// TIA Portal project "ProjectTest" (V15.1)

(* hardware
DEVICE "S7-1200 station_1"  S7-1200 Station
   slot 0: "Rack_0"  S7-1200 Rack  Rack  V1.0
   slot 1: "PLC_1"  CPU 1214C DC/DC/DC  6ES7 214-1AG40-0XB0  V4.2
DEVICE "HMI_1"  KTP900 Basic PN
   slot 0: "HMI_1"  KTP900 Basic PN  6AV2 123-2JB03-0AX0  15.1.0.0
   slot 1: "HMI_RT_1"  KTP900 Basic PN  6AV2 123-2JB03-0AX0  15.1.0.0
   slot 5: "HMI_1.IE_CP_1"  PROFINET Interface  15.0.1.0
      slot 1: "PROFINET Interface_1"  PROFINET Interface
         slot 1: "Port_1"  Port
*)

// ===== PLC "PLC_1"  CPU 1214C DC/DC/DC =====

VAR_GLOBAL   // PLC tag table "Default tag table"
   "System_Byte" AT %MB1 : Byte;
   "FirstScan" AT %M1.0 : Bool;
   "DiagStatusUpdate" AT %M1.1 : Bool;
   "AlwaysTRUE" AT %M1.2 : Bool;
   "AlwaysFALSE" AT %M1.3 : Bool;
   "Clock_Byte" AT %MB0 : Byte;
   "Clock_10Hz" AT %M0.0 : Bool;
   "Clock_5Hz" AT %M0.1 : Bool;
   "Clock_2.5Hz" AT %M0.2 : Bool;
   "Clock_2Hz" AT %M0.3 : Bool;
   "Clock_1.25Hz" AT %M0.4 : Bool;
   "Clock_1Hz" AT %M0.5 : Bool;
   "Clock_0.625Hz" AT %M0.6 : Bool;
   "Clock_0.5Hz" AT %M0.7 : Bool;
   "puls" AT %M2.0 : Bool;
END_VAR

VAR_GLOBAL   // PLC tag table "Tags_DI"
   "Pompa1" AT %Q0.0 : Bool;
   "Pompa2" AT %Q0.1 : Bool;
   "Vana Consum" AT %Q0.2 : Bool;
   "Buton pompa1" AT %I0.0 : Bool;
   "Buton Pompa2" AT %I0.1 : Bool;
   "Buton Vana" AT %I0.2 : Bool;
   "Resetare Contor1" AT %I0.3 : Bool;
   "Resetare Contor2" AT %I0.4 : Bool;
   "Indicatie Pompa1" AT %I0.5 : Bool;
   "Indicatie Pompa2" AT %I0.6 : Bool;
   "Indicatie mod" AT %I0.7 : Bool;
END_VAR

DATA_BLOCK "Bazin"   // DB1
{ S7_Optimized_Access := 'TRUE' }
VERSION : 0.1
   VAR
      Nivel : Real;
      "Vana golire" : Bool := false;
      "Debit golire" : Int := 10;
      Cheie : Int := 1;
      Stare_rising_edge : Bool;
   END_VAR
BEGIN
END_DATA_BLOCK

DATA_BLOCK "Pompa_1"   // DB2
{ S7_Optimized_Access := 'TRUE' }
VERSION : 0.1
   VAR
      Stare : Bool;
      Capacitate : Real := 15.0;
      "Mod" : Int;
      Contor : UInt;
      Stare_rising_edge_bazin : Bool;
      Reset : Bool;
      add_15l : Real := 15.0;
      Stare_rising_edge_pompa : Bool;
   END_VAR
BEGIN
END_DATA_BLOCK

DATA_BLOCK "Pompa_2"   // DB3
{ S7_Optimized_Access := 'TRUE' }
VERSION : 0.1
   VAR
      Stare : Bool;
      Capacitate : Real := 15.0;
      "Mod" : Int;
      Contor : UInt;
      Stare_rising_edge_bazin : Bool;
      Reset : Bool;
      add_15l : Real := 15.0;
      State_rising_edge_pompa : Bool;
   END_VAR
BEGIN
END_DATA_BLOCK

DATA_BLOCK "Adauga  15L la bazin_DB"   // DB4
{ S7_Optimized_Access := 'TRUE' }
VERSION : 0.1
// stored: InstanceOfName Adauga 15L la bazin
"Adauga  15L la bazin"
BEGIN
END_DATA_BLOCK

DATA_BLOCK "Adauga  15L la bazin_DB_1"   // DB5
{ S7_Optimized_Access := 'TRUE' }
VERSION : 0.1
// stored: InstanceOfName Adauga 15L la bazin
"Adauga  15L la bazin"
BEGIN
END_DATA_BLOCK

DATA_BLOCK "Adauga  15L la bazin_DB_2"   // DB6
{ S7_Optimized_Access := 'TRUE' }
VERSION : 0.1
// stored: InstanceOfName Adauga 15L la bazin
"Adauga  15L la bazin"
BEGIN
END_DATA_BLOCK

DATA_BLOCK "Adauga  15L la bazin_DB_3"   // DB7
{ S7_Optimized_Access := 'TRUE' }
VERSION : 0.1
// stored: InstanceOfName Adauga 15L la bazin
"Adauga  15L la bazin"
BEGIN
END_DATA_BLOCK

DATA_BLOCK "Adauga  15L la bazin_DB_4"   // DB8
{ S7_Optimized_Access := 'TRUE' }
VERSION : 0.1
// stored: InstanceOfName Adauga 15L la bazin
"Adauga  15L la bazin"
BEGIN
END_DATA_BLOCK

DATA_BLOCK "Adauga  15L la bazin_DB_5"   // DB9
{ S7_Optimized_Access := 'TRUE' }
VERSION : 0.1
// stored: InstanceOfName Adauga 15L la bazin
"Adauga  15L la bazin"
BEGIN
END_DATA_BLOCK

FUNCTION_BLOCK "Adauga  15L la bazin"   // FB1, LAD
{ S7_Optimized_Access := 'TRUE' }
VERSION : 0.1
   VAR_INPUT
      Input_2 : Bool;
   END_VAR
   VAR_TEMP
      clock_rising_edge : Bool;
   END_VAR
   VAR_TEMP   // added for the SCL form of the ladder/FBD networks
      _w1 : Bool;
      _w2 : Bool;
   END_VAR
BEGIN

REGION Network 1
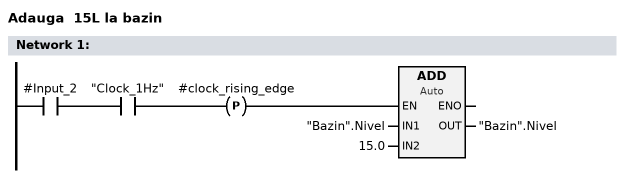
   RUNG wire#powerrail
      Contact( #Input_2 )
      Contact( "Clock_1Hz" )
      P_Trig( #clock_rising_edge )
      Add(in1 := "Bazin".Nivel, in2 := 15.0, out => "Bazin".Nivel)
   END_RUNG
   // the same network as SCL:
   #_w1 := #Input_2 AND "Clock_1Hz";
   #_w2 := #_w1 AND NOT #clock_rising_edge;   // rising edge
   #clock_rising_edge := #_w1;
   IF #_w2 THEN "Bazin".Nivel := "Bazin".Nivel + 15.0; END_IF;
END_REGION
END_FUNCTION_BLOCK

FUNCTION "Block_1" : Void   // FC1, LAD
{ S7_Optimized_Access := 'TRUE' }
VERSION : 0.1
   VAR_INPUT
      input1 : Bool;
   END_VAR
   VAR_TEMP
      clock_rising_edge : Bool;
   END_VAR
   VAR_TEMP   // added for the SCL form of the ladder/FBD networks
      _w1 : Bool;
      _w2 : Bool;
   END_VAR
BEGIN

REGION Network 1
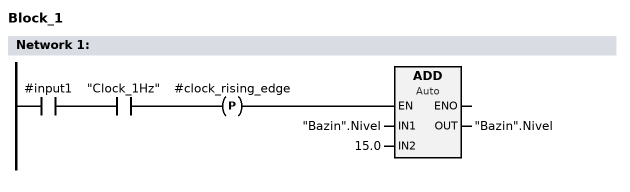
   RUNG wire#powerrail
      Contact( #input1 )
      Contact( "Clock_1Hz" )
      P_Trig( #clock_rising_edge )
      Add(in1 := "Bazin".Nivel, in2 := 15.0, out => "Bazin".Nivel)
   END_RUNG
   // the same network as SCL:
   #_w1 := #input1 AND "Clock_1Hz";
   #_w2 := #_w1 AND NOT #clock_rising_edge;   // rising edge
   #clock_rising_edge := #_w1;
   IF #_w2 THEN "Bazin".Nivel := "Bazin".Nivel + 15.0; END_IF;
END_REGION
END_FUNCTION

ORGANIZATION_BLOCK "Main"   // OB1, LAD, ProgramCycle
TITLE = "Main Program Sweep (Cycle)"
{ S7_Optimized_Access := 'TRUE' }
VERSION : 0.1
   VAR_INPUT
      Initial_Call : Bool;   // Initial call of this OB
      Remanence : Bool;   // =True, if remanent data are available
   END_VAR
   VAR_TEMP   // added for the SCL form of the ladder/FBD networks
      _w1 : Bool;
      _w2 : Bool;
      _w3 : Bool;
      _w4 : Bool;
   END_VAR
BEGIN

REGION Network 1: moduri de functionare
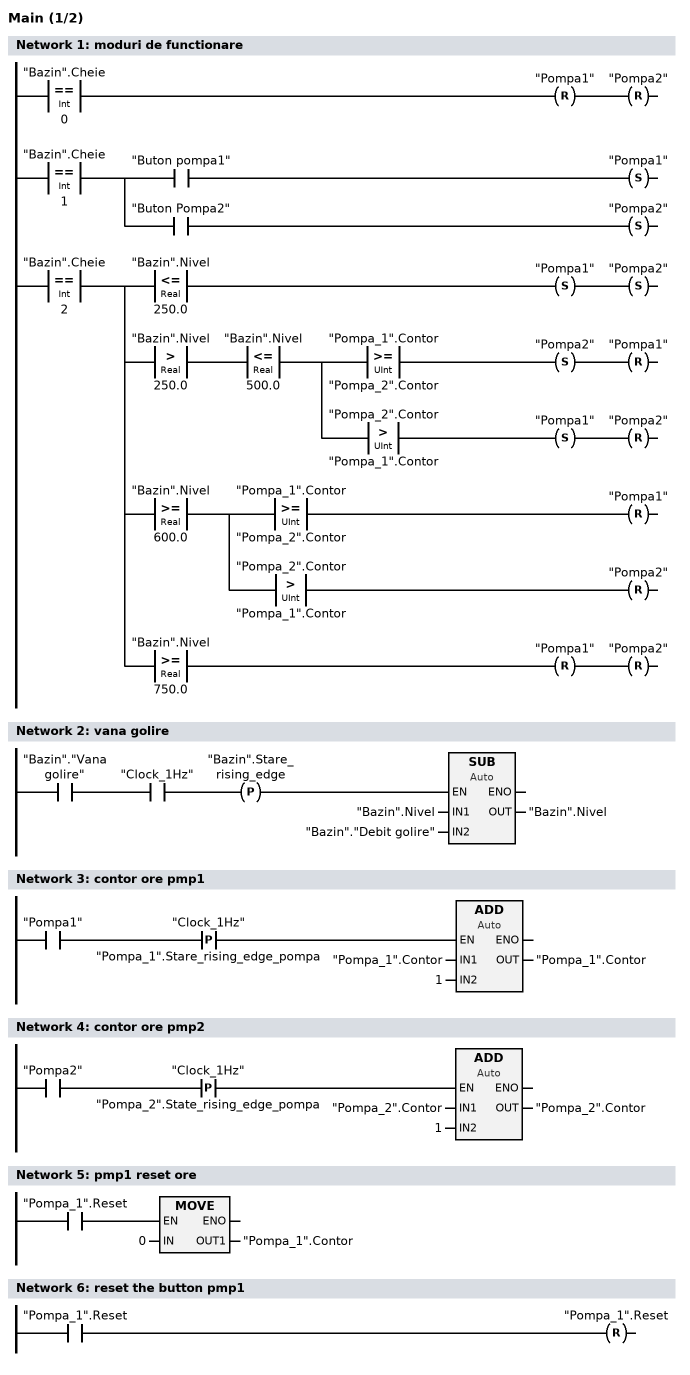
   RUNG wire#powerrail
      { S7_Templates := "SrcType := Int" } EQ_Contact(in1 := "Bazin".Cheie, in2 := 0)
      R_Coil( "Pompa1" )
      R_Coil( "Pompa2" )
   END_RUNG
   RUNG wire#powerrail
      { S7_Templates := "SrcType := Int" } EQ_Contact(in1 := "Bazin".Cheie, in2 := 1)
      wire#w1
      Contact( "Buton pompa1" )
      S_Coil( "Pompa1" )
   END_RUNG
   RUNG wire#w1
      Contact( "Buton Pompa2" )
      S_Coil( "Pompa2" )
   END_RUNG
   RUNG wire#powerrail
      { S7_Templates := "SrcType := Int" } EQ_Contact(in1 := "Bazin".Cheie, in2 := 2)
      wire#w2
      { S7_Templates := "SrcType := Real" } LE_Contact(in1 := "Bazin".Nivel, in2 := 250.0)
      S_Coil( "Pompa1" )
      S_Coil( "Pompa2" )
   END_RUNG
   RUNG wire#w2
      { S7_Templates := "SrcType := Real" } GT_Contact(in1 := "Bazin".Nivel, in2 := 250.0)
      { S7_Templates := "SrcType := Real" } LE_Contact(in1 := "Bazin".Nivel, in2 := 500.0)
      wire#w3
      { S7_Templates := "SrcType := UInt" } GE_Contact(in1 := "Pompa_1".Contor, in2 := "Pompa_2".Contor)
      S_Coil( "Pompa2" )
      R_Coil( "Pompa1" )
   END_RUNG
   RUNG wire#w3
      { S7_Templates := "SrcType := UInt" } GT_Contact(in1 := "Pompa_2".Contor, in2 := "Pompa_1".Contor)
      S_Coil( "Pompa1" )
      R_Coil( "Pompa2" )
   END_RUNG
   RUNG wire#w2
      { S7_Templates := "SrcType := Real" } GE_Contact(in1 := "Bazin".Nivel, in2 := 600.0)
      wire#w4
      { S7_Templates := "SrcType := UInt" } GE_Contact(in1 := "Pompa_1".Contor, in2 := "Pompa_2".Contor)
      R_Coil( "Pompa1" )
   END_RUNG
   RUNG wire#w4
      { S7_Templates := "SrcType := UInt" } GT_Contact(in1 := "Pompa_2".Contor, in2 := "Pompa_1".Contor)
      R_Coil( "Pompa2" )
   END_RUNG
   RUNG wire#w2
      { S7_Templates := "SrcType := Real" } GE_Contact(in1 := "Bazin".Nivel, in2 := 750.0)
      R_Coil( "Pompa1" )
      R_Coil( "Pompa2" )
   END_RUNG
   // the same network as SCL:
   IF "Bazin".Cheie = 0 THEN
       "Pompa1" := FALSE;
       "Pompa2" := FALSE;
   END_IF;
   #_w1 := "Bazin".Cheie = 1;
   IF #_w1 AND "Buton pompa1" THEN "Pompa1" := TRUE; END_IF;
   IF #_w1 AND "Buton Pompa2" THEN "Pompa2" := TRUE; END_IF;
   #_w2 := "Bazin".Cheie = 2;
   IF #_w2 AND ("Bazin".Nivel <= 250.0) THEN
       "Pompa1" := TRUE;
       "Pompa2" := TRUE;
   END_IF;
   #_w3 := #_w2 AND ("Bazin".Nivel > 250.0) AND ("Bazin".Nivel <= 500.0);
   IF #_w3 AND ("Pompa_1".Contor >= "Pompa_2".Contor) THEN
       "Pompa2" := TRUE;
       "Pompa1" := FALSE;
   END_IF;
   IF #_w3 AND ("Pompa_2".Contor > "Pompa_1".Contor) THEN
       "Pompa1" := TRUE;
       "Pompa2" := FALSE;
   END_IF;
   #_w4 := #_w2 AND ("Bazin".Nivel >= 600.0);
   IF #_w4 AND ("Pompa_1".Contor >= "Pompa_2".Contor) THEN "Pompa1" := FALSE; END_IF;
   IF #_w4 AND ("Pompa_2".Contor > "Pompa_1".Contor) THEN "Pompa2" := FALSE; END_IF;
   IF #_w2 AND ("Bazin".Nivel >= 750.0) THEN
       "Pompa1" := FALSE;
       "Pompa2" := FALSE;
   END_IF;
END_REGION

REGION Network 2: vana golire
   RUNG wire#powerrail
      Contact( "Bazin"."Vana golire" )
      Contact( "Clock_1Hz" )
      P_Trig( "Bazin".Stare_rising_edge )
      Sub(in1 := "Bazin".Nivel, in2 := "Bazin"."Debit golire", out => "Bazin".Nivel)
   END_RUNG
   // the same network as SCL:
   #_w1 := "Bazin"."Vana golire" AND "Clock_1Hz";
   #_w2 := #_w1 AND NOT "Bazin".Stare_rising_edge;   // rising edge
   "Bazin".Stare_rising_edge := #_w1;
   IF #_w2 THEN "Bazin".Nivel := "Bazin".Nivel - "Bazin"."Debit golire"; END_IF;
END_REGION

REGION Network 3: contor ore pmp1
   RUNG wire#powerrail
      Contact( "Pompa1" )
      P_Contact(operand := "Clock_1Hz", bit := "Pompa_1".Stare_rising_edge_pompa)
      Add(in1 := "Pompa_1".Contor, in2 := 1, out => "Pompa_1".Contor)
   END_RUNG
   // the same network as SCL:
   #_w1 := "Pompa1" AND "Clock_1Hz" AND NOT "Pompa_1".Stare_rising_edge_pompa;   // rising edge of "Clock_1Hz"
   "Pompa_1".Stare_rising_edge_pompa := "Clock_1Hz";
   IF #_w1 THEN "Pompa_1".Contor := "Pompa_1".Contor + 1; END_IF;
END_REGION

REGION Network 4: contor ore pmp2
   RUNG wire#powerrail
      Contact( "Pompa2" )
      P_Contact(operand := "Clock_1Hz", bit := "Pompa_2".State_rising_edge_pompa)
      Add(in1 := "Pompa_2".Contor, in2 := 1, out => "Pompa_2".Contor)
   END_RUNG
   // the same network as SCL:
   #_w1 := "Pompa2" AND "Clock_1Hz" AND NOT "Pompa_2".State_rising_edge_pompa;   // rising edge of "Clock_1Hz"
   "Pompa_2".State_rising_edge_pompa := "Clock_1Hz";
   IF #_w1 THEN "Pompa_2".Contor := "Pompa_2".Contor + 1; END_IF;
END_REGION

REGION Network 5: pmp1 reset ore
   RUNG wire#powerrail
      Contact( "Pompa_1".Reset )
      Move(in := 0, out1 => "Pompa_1".Contor)
   END_RUNG
   // the same network as SCL:
   IF "Pompa_1".Reset THEN "Pompa_1".Contor := 0; END_IF;
END_REGION

REGION Network 6: reset the button pmp1
   RUNG wire#powerrail
      Contact( "Pompa_1".Reset )
      R_Coil( "Pompa_1".Reset )
   END_RUNG
   // the same network as SCL:
   IF "Pompa_1".Reset THEN "Pompa_1".Reset := FALSE; END_IF;
END_REGION

REGION Network 7: pmp 2 reset ore
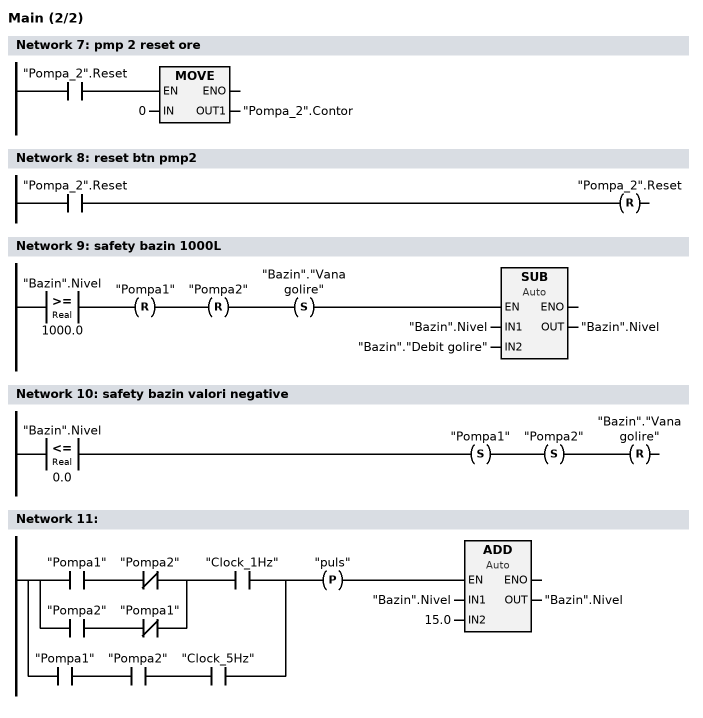
   RUNG wire#powerrail
      Contact( "Pompa_2".Reset )
      Move(in := 0, out1 => "Pompa_2".Contor)
   END_RUNG
   // the same network as SCL:
   IF "Pompa_2".Reset THEN "Pompa_2".Contor := 0; END_IF;
END_REGION

REGION Network 8: reset btn pmp2
   RUNG wire#powerrail
      Contact( "Pompa_2".Reset )
      R_Coil( "Pompa_2".Reset )
   END_RUNG
   // the same network as SCL:
   IF "Pompa_2".Reset THEN "Pompa_2".Reset := FALSE; END_IF;
END_REGION

REGION Network 9: safety bazin 1000L
   RUNG wire#powerrail
      { S7_Templates := "SrcType := Real" } GE_Contact(in1 := "Bazin".Nivel, in2 := 1000.0)
      R_Coil( "Pompa1" )
      R_Coil( "Pompa2" )
      S_Coil( "Bazin"."Vana golire" )
      Sub(in1 := "Bazin".Nivel, in2 := "Bazin"."Debit golire", out => "Bazin".Nivel)
   END_RUNG
   // the same network as SCL:
   IF "Bazin".Nivel >= 1000.0 THEN
       "Pompa1" := FALSE;
       "Pompa2" := FALSE;
       "Bazin"."Vana golire" := TRUE;
       "Bazin".Nivel := "Bazin".Nivel - "Bazin"."Debit golire";
   END_IF;
END_REGION

REGION Network 10: safety bazin valori negative
   RUNG wire#powerrail
      { S7_Templates := "SrcType := Real" } LE_Contact(in1 := "Bazin".Nivel, in2 := 0.0)
      S_Coil( "Pompa1" )
      S_Coil( "Pompa2" )
      R_Coil( "Bazin"."Vana golire" )
   END_RUNG
   // the same network as SCL:
   IF "Bazin".Nivel <= 0.0 THEN
       "Pompa1" := TRUE;
       "Pompa2" := TRUE;
       "Bazin"."Vana golire" := FALSE;
   END_IF;
END_REGION

REGION Network 11
   RUNG wire#powerrail
      Contact( "Pompa1" )
      I_Contact( "Pompa2" )
      wire#w1
      Contact( "Clock_1Hz" )
      wire#w2
      P_Trig( "puls" )
      Add(in1 := "Bazin".Nivel, in2 := 15.0, out => "Bazin".Nivel)
   END_RUNG
   RUNG wire#powerrail
      Contact( "Pompa2" )
      I_Contact( "Pompa1" )
   END_RUNG wire#w1
   RUNG wire#powerrail
      Contact( "Pompa1" )
      Contact( "Pompa2" )
      Contact( "Clock_5Hz" )
   END_RUNG wire#w2
   // the same network as SCL:
   #_w1 := ((("Pompa1" AND NOT "Pompa2") OR ("Pompa2" AND NOT "Pompa1")) AND "Clock_1Hz") OR ("Pompa1" AND "Pompa2" AND "Clock_5Hz");
   #_w2 := #_w1 AND NOT "puls";   // rising edge
   "puls" := #_w1;
   IF #_w2 THEN "Bazin".Nivel := "Bazin".Nivel + 15.0; END_IF;
END_REGION
END_ORGANIZATION_BLOCK

(* ===== HMI "HMI_RT_1" =====
system functions are stored by id; their names below are inferred from use
connection "HMI_Connection_1": ETHERNET, SMART_S7_1200_OMS

HMI tags "Default tag table"
   "Bazin_Nivel" : Real = PLC Bazin.Nivel, 1 s
   "Bazin_Vana golire" : Bool = PLC Bazin."Vana golire", 1 s
   "Pompa_1_Contor" : UInt = PLC Pompa_1.Contor, 1 s
   "Pompa_2_Contor" : UInt = PLC Pompa_2.Contor, 1 s
   "Pompa_1_Reset" : Bool = PLC Pompa_1.Reset, 1 s
   "Pompa_2_Reset" : Bool = PLC Pompa_2.Reset, 1 s
   "Bazin_Cheie" : Int = PLC Bazin.Cheie, 1 s
   "Pompa1" : Bool = PLC Pompa1 AT %Q0.0, 1 s
   "Pompa2" : Bool = PLC Pompa2 AT %Q0.1, 1 s

screen "Screen_1" 800x480
   Bar "Bar_1" at 259,52 size 164x377; MinimumValue 0; MaximumValue 1000
      ProcessValue <- "Bazin_Nivel"
   Button "Button_1" at 85,411 size 96x32; TextOff 'Reset vana'
      on Click: SetBit("Bazin_Vana golire")
   IOField "I/O field_1" at 480,77 size 96x32; FormatPattern 99999; Unit s
      ProcessValue <- "Pompa_1_Contor"
   TextField "Text field_1" at 480,53 size 96x20; Text 'Counter pmp1'
   IOField "I/O field_2" at 486,154 size 96x32; FormatPattern 99999; Unit s
      ProcessValue <- "Pompa_2_Contor"
   TextField "Text field_2" at 486,134 size 96x20; Text 'Counter pmp2'
   Button "Button_2" at 610,78 size 96x32; TextOff 'Reset1'
      on Click: SetBit("Pompa_1_Reset")
   Button "Button_3" at 609,153 size 96x32; TextOff 'Reset2'
      on Activate: SetBit("Pompa_2_Reset")
   Button "Button_4" at 56,117 size 96x32; TextOff '0'
      on Click: SetTag("Bazin_Cheie", 0)
   Button "Button_5" at 56,185 size 96x32; TextOff '1'
      on Click: SetTag("Bazin_Cheie", 1)
   Button "Button_6" at 56,250 size 96x32; TextOff '2'
      on Click: SetTag("Bazin_Cheie", 2)
   TextField "Text field_3" at 65,67 size 70x20; Text 'Set config'
   Rectangle "Rectangle_1" at 85,351 size 96x48
      Appearance <- "Bazin_Vana golire"
   Circle "Circle_1" at 505,319 size 48x48
      Appearance <- "Pompa1"
   Circle "Circle_2" at 593,321 size 48x48
      Appearance <- "Pompa2"
   TextField "Text field_4" at 505,299 size 40x20; Text 'Pmp1'
   TextField "Text field_5" at 593,302 size 40x20; Text 'Pmp2'
   Button "Button_7" at 610,223 size 96x32; TextOff 'doar reset'
*)